// TIA Portal project "TESTV18" (V18)

(* hardware
DEVICE "Stazione S7-1500/ET200MP_1"  S7-1500 station
   slot 0: "Telaio di montaggio_0"  Rack  6ES7 590-1***0-0AA0
   slot 1: "PLC"  CPU 1511F-1 PN  6ES7 511-1FK02-0AB0  V2.8
      slot 3: "Display CPU_1"  6ES7591-1AA00-0AA0
      slot 32768: "Interfaccia PROFINET_1"  X1
         slot 32769: "Porta_1"  X1 P1
         slot 32770: "Porta_2"  X1 P2
      slot 34817: "Virtual CP interface port_1"  Virtual CP interface port  Virtual CP interface port
   slot 2: "AQ 4xU/I ST_1"  AQ 4xU/I ST  6ES7 532-5HD00-0AB0  V2.0
   slot 3: "AI 8xU/I HS_1"  AI 8xU/I HS  6ES7 531-7NF10-0AB0  V2.0
   slot 4: "DI 16x24VDC HF_1"  DI 16x24VDC HF  6ES7 521-1BH00-0AB0  V2.0
   slot 5: "DQ 16x24VDC/0.5A ST_1"  DQ 16x24VDC/0.5A ST  6ES7 522-1BH00-0AB0  V2.0
DEVICE "HMI"  TP700 Comfort
   slot 0: "HMI"  TP700 Comfort  6AV2 124-0GC01-0AX0  17.0.0.0
   slot 1: "HMI_RT_1"  TP700 Comfort  6AV2 124-0GC01-0AX0  17.0.0.0
   slot 5: "HMI.IE_CP_1"  PROFINET Interface  17.0.0.0
      slot 1: "Interfaccia_1 PROFINET"  PROFINET Interface
         slot 1: "Porta_1"  Port
         slot 2: "Porta_2"  Port
   slot 7: "HMI.MPI/DP_CP_1"  MPI/DP Interface  17.0.0.0
DEVICE "GSD device_1"  GSD.Device.PN
   slot 0: "Telaio di montaggio"  Rack  V1.0
   slot 0: "IAIPRT1"  RT Standard  IAI-PRT
      slot 0: "RT Standard"  RT Standard
      slot 1: "Interface"  Interface
         slot 1: "Port 1"  Port 1
   slot 1: "Input 1 word_1"  Input 1 word  IAI-PRT
      slot 0: "Input 1 word"  Input 1 word
   slot 2: "Input 1 word_2"  Input 1 word  IAI-PRT
      slot 0: "Input 1 word"  Input 1 word
   slot 3: "Input 1 word_3"  Input 1 word  IAI-PRT
      slot 0: "Input 1 word"  Input 1 word
   slot 4: "Input 1 word_4"  Input 1 word  IAI-PRT
      slot 0: "Input 1 word"  Input 1 word
   slot 5: "Input 1 word_5"  Input 1 word  IAI-PRT
      slot 0: "Input 1 word"  Input 1 word
   slot 6: "Input 1 word_6"  Input 1 word  IAI-PRT
      slot 0: "Input 1 word"  Input 1 word
   slot 7: "Input 1 word_7"  Input 1 word  IAI-PRT
      slot 0: "Input 1 word"  Input 1 word
   slot 8: "Input 1 word_8"  Input 1 word  IAI-PRT
      slot 0: "Input 1 word"  Input 1 word
   slot 9: "Input 1 word_9"  Input 1 word  IAI-PRT
      slot 0: "Input 1 word"  Input 1 word
   slot 10: "Input 1 word_10"  Input 1 word  IAI-PRT
      slot 0: "Input 1 word"  Input 1 word
   slot 11: "Input 1 word_11"  Input 1 word  IAI-PRT
      slot 0: "Input 1 word"  Input 1 word
   slot 12: "Input 1 word_12"  Input 1 word  IAI-PRT
      slot 0: "Input 1 word"  Input 1 word
   slot 13: "Input 1 word_13"  Input 1 word  IAI-PRT
      slot 0: "Input 1 word"  Input 1 word
   slot 14: "Input 1 word_14"  Input 1 word  IAI-PRT
      slot 0: "Input 1 word"  Input 1 word
   slot 15: "Input 1 word_15"  Input 1 word  IAI-PRT
      slot 0: "Input 1 word"  Input 1 word
   slot 16: "Input 1 word_16"  Input 1 word  IAI-PRT
      slot 0: "Input 1 word"  Input 1 word
   slot 17: "Output 1 word_1"  Output 1 word  IAI-PRT
      slot 0: "Output 1 word"  Output 1 word
   slot 18: "Output 1 word_2"  Output 1 word  IAI-PRT
      slot 0: "Output 1 word"  Output 1 word
   slot 19: "Output 1 word_3"  Output 1 word  IAI-PRT
      slot 0: "Output 1 word"  Output 1 word
   slot 20: "Output 1 word_4"  Output 1 word  IAI-PRT
      slot 0: "Output 1 word"  Output 1 word
   slot 21: "Output 1 word_5"  Output 1 word  IAI-PRT
      slot 0: "Output 1 word"  Output 1 word
   slot 22: "Output 1 word_6"  Output 1 word  IAI-PRT
      slot 0: "Output 1 word"  Output 1 word
   slot 23: "Output 1 word_7"  Output 1 word  IAI-PRT
      slot 0: "Output 1 word"  Output 1 word
   slot 24: "Output 1 word_8"  Output 1 word  IAI-PRT
      slot 0: "Output 1 word"  Output 1 word
   slot 25: "Output 1 word_9"  Output 1 word  IAI-PRT
      slot 0: "Output 1 word"  Output 1 word
   slot 26: "Output 1 word_10"  Output 1 word  IAI-PRT
      slot 0: "Output 1 word"  Output 1 word
   slot 27: "Output 1 word_11"  Output 1 word  IAI-PRT
      slot 0: "Output 1 word"  Output 1 word
   slot 28: "Output 1 word_12"  Output 1 word  IAI-PRT
      slot 0: "Output 1 word"  Output 1 word
   slot 29: "Output 1 word_13"  Output 1 word  IAI-PRT
      slot 0: "Output 1 word"  Output 1 word
   slot 30: "Output 1 word_14"  Output 1 word  IAI-PRT
      slot 0: "Output 1 word"  Output 1 word
   slot 31: "Output 1 word_15"  Output 1 word  IAI-PRT
      slot 0: "Output 1 word"  Output 1 word
   slot 32: "Output 1 word_16"  Output 1 word  IAI-PRT
      slot 0: "Output 1 word"  Output 1 word
*)

// ===== PLC "PLC"  CPU 1511F-1 PN =====

VAR_GLOBAL   // PLC tag table "Tabella delle variabili standard"
   "System_Byte" AT %MB16382 : Byte;
   "FirstScan" AT %M16382.0 : Bool;
   "DiagStatusUpdate" AT %M16382.1 : Bool;
   "AlwaysTRUE" AT %M16382.2 : Bool;
   "AlwaysFALSE" AT %M16382.3 : Bool;
   "Clock_Byte" AT %MB16383 : Byte;
   "Clock_10Hz" AT %M16383.0 : Bool;
   "Clock_5Hz" AT %M16383.1 : Bool;
   "Clock_2.5Hz" AT %M16383.2 : Bool;
   "Clock_2Hz" AT %M16383.3 : Bool;
   "Clock_1.25Hz" AT %M16383.4 : Bool;
   "Clock_1Hz" AT %M16383.5 : Bool;
   "Clock_0.625Hz" AT %M16383.6 : Bool;
   "Clock_0.5Hz" AT %M16383.7 : Bool;
   "Tag_1" AT %M0.0 : Bool;
   "Tag_2" AT %M0.1 : Bool;
   "Tag_3" AT %M0.3 : Bool;
   "Tag_4" AT %M0.4 : Bool;
   "Tag_5" AT %M0.5 : Bool;
   "Tag_6" AT %M0.6 : Bool;
   "Tag_7" AT %M0.7 : Bool;
   "Tag_8" AT %M500.0 : Bool;
   "Tag_9" AT %T100 : Timer;
   "Tag_10" AT %M0.2 : Bool;
   "Tag_11" AT %M2.0 : Bool;
   "Tag_12" AT %MD1000 : DWord;
   "Tag_13" AT %MW1000 : Word;
   "Tag_14" AT %MW1004 : UInt;
   "Tag_15" AT %Q2.0 : Bool;
   "Tag_16" AT %M5.0 : Bool;
   "Tag_17" AT %M5.1 : Bool;
   "Tag_18" AT %M5.2 : Bool;
   "Tag_19" AT %M5.3 : Bool;
   "Tag_20" AT %M4.0 : Bool;
   "Tag_21" AT %M4.1 : Bool;
   "Tag_22" AT %M3.0 : Bool;
   "Tag_23" AT %IW0 : Word;
   "Tag_24" AT %IB0 : Byte;
   "Tag_25" AT %IB16 : Byte;
   "Tag_26" AT %M2.1 : Bool;
   "Tag_27" AT %M2.3 : Bool;
   "Tag_28" AT %M2.4 : Bool;
   "Tag_29" AT %M2.5 : Bool;
   "Tag_30" AT %M2.6 : Bool;
   "Tag_31" AT %M2.7 : Bool;
   "Tag_32" AT %M2.2 : Bool;
   "Tag_33" AT %M3.1 : Bool;
   "Tag_34" AT %M3.2 : Bool;
   "Tag_35" AT %Q9.7 : Bool;
   "TGT_Pos" AT %QD10 : DWord;   // Position to be reached
   "Tag_37" AT %QD13 : DWord;
   "Tag_38" AT %QW10 : Word;
   "Tag_39" AT %QW11 : Word;
   "Tag_40" AT %QW13 : Word;
   "Tag_41" AT %QD12 : DWord;
   "Tag_42" AT %QD11 : DWord;
   "Tag_43" AT %QD34 : DWord;
   "CTRL_Sig2" AT %QD38 : DWord;   // Control dword signal 2
   "POS_BAND" AT %QD14 : DWord;   // Positioning band
   "SPE_mms" AT %QD18 : DWord;   // Speed mm/s
   "ZBO_ZBP" AT %QD22 : DWord;   // Zone boundary+
   "ZBO_ZBM" AT %QD26 : DWord;   // Zone boundary-
   "ACC_Accell" AT %QW30 : Word;   // Acceleration
   "DCL_Decell" AT %QW32 : Word;   // Deceleration
   "PLV_PressLimV" AT %QW34 : Word;   // Pressing current-limiting value
   "LCT_LoadCurrTh" AT %QW36 : Word;   // Load current threshold
   "Tag_36" AT %M1.0 : Bool;
   "Curr_POS" AT %ID18 : DWord;   // Current Position
   "Curr_CMD" AT %ID22 : DInt;   // Current command
   "Curr_SPD" AT %ID26 : UDInt;   // Current Speed
   "Allarm_COD" AT %ID30 : UDInt;   // Allarm Code
   "TotalMove_CNT" AT %ID38 : DInt;   // Total moving counter
   "TotalMove_DST" AT %ID42 : UDInt;   // Total moving distance
   "Status_DW" AT %ID46 : DWord;   // Status words PCON->PLC
END_VAR

TYPE "IAI_PCONPRTFM32OUT"
TITLE = IAI_PCONPRTFM32OUT
// Data type used for IAI PCON controller profinet configured in full mode (3 on parameter 84) with 32 word I/O occupied (0 on parameter 90)
   STRUCT
      Target_POS : DInt;   // Set the target position on the absolute coordinates.
      Positioning_BAND : UDInt;   // Positioning band
      Speed : UDInt;   // Specify the speed at which to move the actuator
      ZoneBNDP_BNDM : UDInt;   // The status signal PZONE turns ON when the current position is inside these +/- boundaries.
      Acceleration : USInt;   // Specify the acceleration at which to move the actuator
      Deceleration : USInt;   // Specify the deceleration at which to move the actuator
      Pressing_CLV : USInt;   // Specify the current- limiting value to be used during pressing operation.
      Load_current_threshold : USInt;   // Set the current threshold in this register when whether or not the load current exceeds the threshold is judged.
      CTRL1 : Struct   // Control WORD 1
         CTRL1_Sig_15 : Bool;   // Unavailable
         CTRL1_Sig_14 : Bool;   // Unavailable
         CTRL1_Sig_NTC1 : Bool;   // NTC1 (ACON only)
         CTRL1_Sig_NTC0 : Bool;   // NTC0 (ACON only)
         CTRL1_Sig_11 : Bool;   // Unavailable
         CTRL1_Sig_SMOD : Bool;   // SMOD (PCON only) Stopping control mode: When this signal is ON, servo control is performed during stopping.
         CTRL1_Sig_ASO1 : Bool;   // ASO1 Stop Mode 1 Select stop mode while standing
         CTRL1_Sig_ASO0 : Bool;   // ASO1 Stop Mode 0 Select stop mode while standing
         CTRL1_Sig_MOD1 : Bool;   // Acceleration / deceleration mode
         CTRL1_Sig_MOD0 : Bool;   // Acceleration / deceleration mode
         CTRL1_Sig_GSL1 : Bool;   // GSL1 (ACON only)
         CTRL1_Sig_GSL0 : Bool;   // GSL0 (ACON only)
         CTRL1_Sig_INC : Bool;   // Incremental Command: Absolute position commands are issued when this signal is OFF
         CTRL1_Sig_DIR : Bool;   // Pressing direction specification: “OFF” for the direction reducing the positioning band from the target position
         CTRL1_Sig_PUSH : Bool;   // Pressing specification : Positioning operation is performed when this signal is OFF
         CTRL1_Sig_00 : Bool;   // Unavailable
      END_STRUCT;
      CTRL2 : Struct   // Control WORD 2
         CTRL2_Sig_BKRL : Bool;   // Forced brake release: When it is turned ON, the brake is released
         CTRL2_Sig_RMOD : Bool;   // Operating mode selector : The AUTO mode is selected when this signal is OFF
         CTRL2_Sig_13 : Bool;   // Unavailable
         CTRL2_Sig_12 : Bool;   // Unavailable
         CTRL2_Sig_11 : Bool;   // Unavailable
         CTRL2_Sig_10 : Bool;   // Unavailable
         CTRL2_Sig_CLBR : Bool;   // Load cell calibration command (Dedicated for PCON-CBP/CGBP)
         "CTRL2_Sig_JOG+" : Bool;   // +Jog: “ON” for Movement in the Opposite Direction of Home
         "CTRL2_Sig_JOG-" : Bool;   // -Jog: “ON” for Movement in the Home Direction
         CTRL2_Sig_JVEL : Bool;   // Jog-speed/inch-distance switching
         CTRL2_Sig_JISL : Bool;   // Jog/inch switching: Jog operation is performed when this signal is OFF
         CTRL2_Sig_SON : Bool;   // GSL0 (ACON only)
         CTRL2_Sig_RES : Bool;   // Reset: A reset is performed when this signal turns ON.
         CTRL2_Sig_STP : Bool;   // Pause: A pause command is issued when this signal turns ON.
         CTRL2_Sig_HOME : Bool;   // Home return: A home-return command is issued when this signal turns ON.
         CTRL2_Sig_DSTR : Bool;   // Positioning start: A move command is issued when this signal turns ON.
      END_STRUCT;
   END_STRUCT;
END_TYPE

TYPE "IAI_PCONPRT"
   STRUCT
      PLCToPCON : "IAI_PCONPRTFM32OUT";
      PCONToPLC : "IAI_PCONPRTFM32IN";
   END_STRUCT;
END_TYPE

TYPE "IAI_PCONPRTFM32IN"
TITLE = IAI_PCONPRTFM32OUT
// Data type used for IAI PCON controller profinet configured in full mode (3 on parameter 84) with 32 word I/O occupied (0 on parameter 90)
   STRUCT
      Current_POS : DInt;   // Stores the current position. The unit is 0.01mm.
      Command_CUR : UDInt;   // Stores the currently commanded current. The unit is mA.
      Current_SPD : DInt;   // The current speed is indicated. The unit is 0.01mm/s. Positive value: The actuator is moving in the direction opposite home.
      Alarm_COD : UDInt;   // Stores an alarm code when an alarm (all alarms including message level ones) is generated.
      Current_LOA : DInt;   // Current load (Dedicated for PCON-CBP /CGBP)The unit is 0.01N.
      TotalMove_CNT : UDInt;   // Total moving conts (unit: times)
      TotalMove_DST : USInt;   // Total moving distance (unit: m)
      CTRL1 : Struct   // Control WORD 1
         STAT1_Sig_15 : Bool;   // Unavailable
         STAT1_Sig_14 : Bool;   // Unavailable
         STAT1_Sig_13 : Bool;   // Unavailable
         STAT1_Sig_12 : Bool;   // Unavailable
         STAT1_Sig_11 : Bool;   // Unavailable
         STAT1_Sig_10 : Bool;   // Unavailable
         STAT1_Sig_09 : Bool;   // Unavailable
         STAT1_Sig_08 : Bool;   // Unavailable
         STAT1_Sig_07 : Bool;   // Unavailable
         STAT1_Sig_06 : Bool;   // Unavailable
         STAT1_Sig_05 : Bool;   // Unavailable
         STAT1_Sig_04 : Bool;   // Unavailable
         STAT1_Sig_03 : Bool;   // Unavailable
         STAT1_Sig_02 : Bool;   // Unavailable
         CTRL1_Sig_CEND : Bool;   // Load cell calibration command. (Dedicated for PCON-CBP/CGBP)
         CTRL1_Sig_ALML : Bool;   // Light error status: Turns ON when light alarm (threshold exceeded for number of movement, etc.) that the operation can be continued with is issued. Note: ALM LED would not turn ON with a light error.
      END_STRUCT;
      CTRL2 : Struct   // Control WORD 2
         CTRL2_Sig_EMGS : Bool;   // Emergency stop: An emergency stop is actuated when this signal turns ON.
         CTRL2_Sig_PWR : Bool;   // Controller ready : This signal turns ON when the controller becomes ready.
         CTRL2_Sig_ZONE2 : Bool;   // Zone 2:“ON” for the current position within the zone set range
         CTRL2_Sig_ZONE1 : Bool;   // Zone 1:“ON” for the current position within the zone set range
         CTRL2_Sig_PZONE : Bool;   // Position zone: This signal turns ON when the current position is inside the specified position zone.
         CTRL2_Sig_LOAD : Bool;   // Load output judgment: When this signal is ON, the specified load has been reached.
         CTRL2_Sig_TRQS : Bool;   // Torque level: When this signal is ON, the specified load has been reached.
         CTRL2_Sig_RMDS : Bool;   // Operation mode status: This signal is OFF when the current mode is AUTO, or ON when the current mode is MANU.
         CTRL2_Sig_GHMS : Bool;   // Under Home return Operation: This signal remains ON while home return is in progress.
         CTRL2_Sig_PUSHS : Bool;   // Pressing in progress: This signal remains ON while pressing operation is in progress.
         CTRL2_Sig_PSFL : Bool;   // Pressing and a Miss: This signal turns ON when the actuator missed the work part in pressing operation.
         CTRL2_Sig_SV : Bool;   // Operation preparation end: This signal turns ON when the servo turns ON.
         CTRL2_Sig_ALM : Bool;   // Alarm: This signal turns ON when an alarm occurs.
         CTRL2_Sig_MOVE : Bool;   // Moving signal: This signal remains ON while the actuator is moving.
         CTRL2_Sig_HEND : Bool;   // Home return completion: This signal turns ON when home return is completed
         CTRL2_Sig_PEND : Bool;   // Positioning completion signal: This signal turns ON when positioning is completed.
      END_STRUCT;
   END_STRUCT;
END_TYPE

DATA_BLOCK "Main_Safety_RTG1_DB"   // DB1, F_DB
{ S7_Optimized_Access := 'TRUE' }
NAME : FUSI
VERSION : 0.1
// stored: InstanceOfName Main_Safety_RTG1
"Main_Safety_RTG1"
BEGIN
END_DATA_BLOCK

DATA_BLOCK "DB_AUX"   // DB3
{ S7_Optimized_Access := 'TRUE' }
VERSION : 0.1
   VAR
      FP : Array[0..10] of Bool;
      TARGET_POS : Array[0..4] of DInt;
      SPEED_POS : Array[0..4] of UDInt;
      ACC_DEC : USInt;
      AXIS1 : "IAI_PCONPRT";
      HMI_Bit : Struct
         HMIb1 : Bool;   // Load POS1
         HMIb2 : Bool;   // Load POS2
         HMIb3 : Bool;   // Load POS3
         HMIb4 : Bool;   // Load POS4
         HMIb5 : Bool;   // Servo ON
         HMIb6 : Bool;   // Start positioning
         HMIb7 : Bool;   // Homing
         HMIb8 : Bool;   // JOG+
         HMIb9 : Bool;   // JOG-
         HMIb10 : Bool;   // Reset allarm
         HMIb11 : Bool;
         HMIb12 : Bool;
         HMIb13 : Bool;
      END_STRUCT;
   END_VAR
BEGIN
END_DATA_BLOCK

FUNCTION_BLOCK "Main_Safety_RTG1"   // FB1, F_FBD
{ S7_Optimized_Access := 'TRUE' }
BEGIN
END_FUNCTION_BLOCK

ORGANIZATION_BLOCK "Main"   // OB1, LAD, ProgramCycle
TITLE = "Main Program Sweep (Cycle)"
{ S7_Optimized_Access := 'TRUE' }
VERSION : 0.1
   VAR_INPUT
      Initial_Call : Bool;   // Initial call of this OB
      Remanence : Bool;   // =True, if remanent data are available
   END_VAR
BEGIN

REGION Network 1: IAI controllers side input register PLC -> PCON
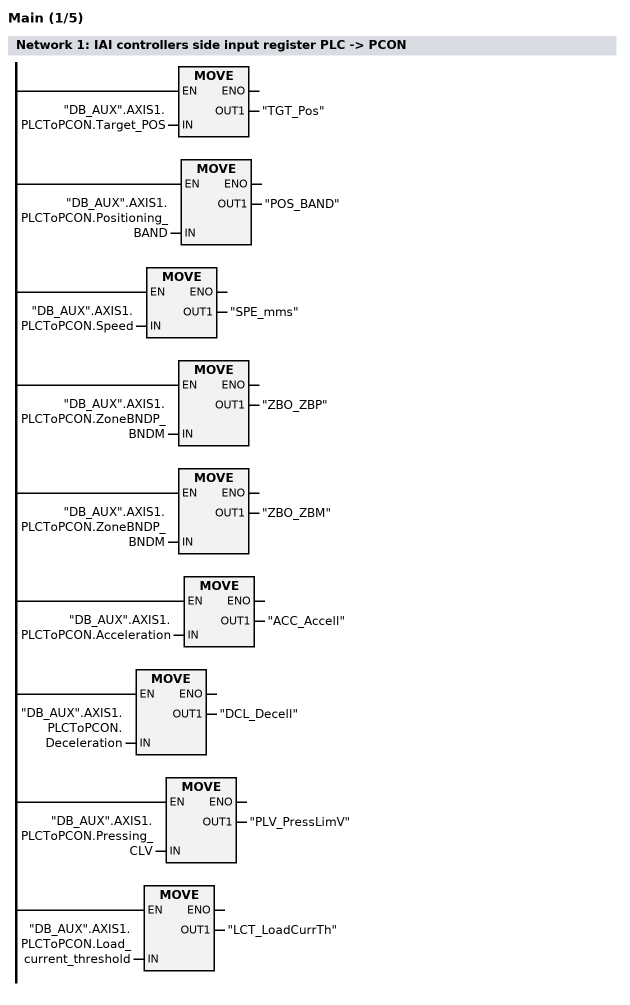
   RUNG wire#powerrail
      Move(in := "DB_AUX".AXIS1.PLCToPCON.Target_POS, out1 => "TGT_Pos")
   END_RUNG
   RUNG wire#powerrail
      Move(in := "DB_AUX".AXIS1.PLCToPCON.Positioning_BAND, out1 => "POS_BAND")
   END_RUNG
   RUNG wire#powerrail
      Move(in := "DB_AUX".AXIS1.PLCToPCON.Speed, out1 => "SPE_mms")
   END_RUNG
   RUNG wire#powerrail
      Move(in := "DB_AUX".AXIS1.PLCToPCON.ZoneBNDP_BNDM, out1 => "ZBO_ZBP")
   END_RUNG
   RUNG wire#powerrail
      Move(in := "DB_AUX".AXIS1.PLCToPCON.ZoneBNDP_BNDM, out1 => "ZBO_ZBM")
   END_RUNG
   RUNG wire#powerrail
      Move(in := "DB_AUX".AXIS1.PLCToPCON.Acceleration, out1 => "ACC_Accell")
   END_RUNG
   RUNG wire#powerrail
      Move(in := "DB_AUX".AXIS1.PLCToPCON.Deceleration, out1 => "DCL_Decell")
   END_RUNG
   RUNG wire#powerrail
      Move(in := "DB_AUX".AXIS1.PLCToPCON.Pressing_CLV, out1 => "PLV_PressLimV")
   END_RUNG
   RUNG wire#powerrail
      Move(in := "DB_AUX".AXIS1.PLCToPCON.Load_current_threshold, out1 => "LCT_LoadCurrTh")
   END_RUNG
   // the same network as SCL:
   "TGT_Pos" := "DB_AUX".AXIS1.PLCToPCON.Target_POS;
   "POS_BAND" := "DB_AUX".AXIS1.PLCToPCON.Positioning_BAND;
   "SPE_mms" := "DB_AUX".AXIS1.PLCToPCON.Speed;
   "ZBO_ZBP" := "DB_AUX".AXIS1.PLCToPCON.ZoneBNDP_BNDM;
   "ZBO_ZBM" := "DB_AUX".AXIS1.PLCToPCON.ZoneBNDP_BNDM;
   "ACC_Accell" := "DB_AUX".AXIS1.PLCToPCON.Acceleration;
   "DCL_Decell" := "DB_AUX".AXIS1.PLCToPCON.Deceleration;
   "PLV_PressLimV" := "DB_AUX".AXIS1.PLCToPCON.Pressing_CLV;
   "LCT_LoadCurrTh" := "DB_AUX".AXIS1.PLCToPCON.Load_current_threshold;
END_REGION

REGION Network 2: IAI controllers side input register PLC -> PCON
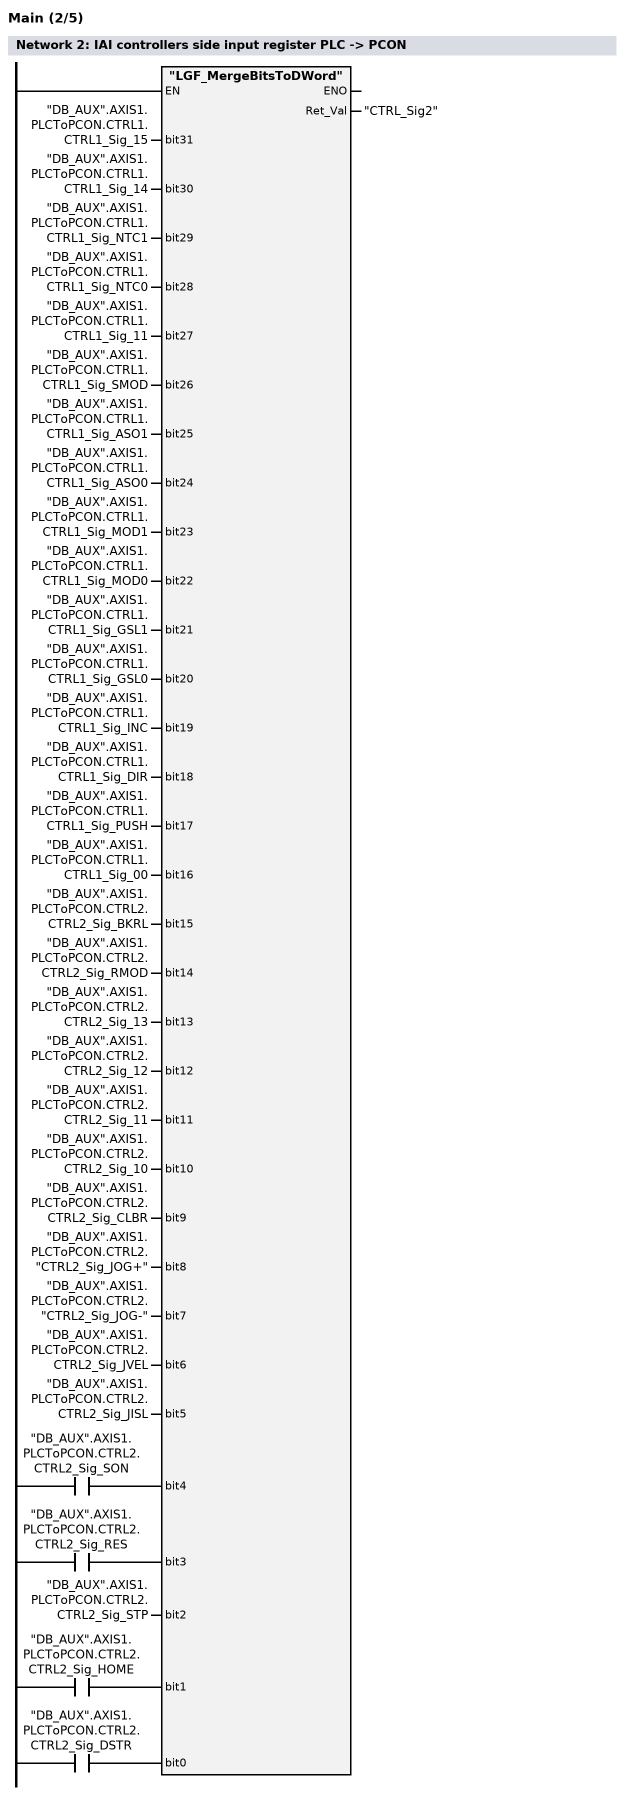
   RUNG wire#powerrail
      "LGF_MergeBitsToDWord"(bit4 := wire#w1, bit3 := wire#w2, bit1 := wire#w3, bit0 := wire#w4, bit31 := "DB_AUX".AXIS1.PLCToPCON.CTRL1.CTRL1_Sig_15, bit30 := "DB_AUX".AXIS1.PLCToPCON.CTRL1.CTRL1_Sig_14, bit29 := "DB_AUX".AXIS1.PLCToPCON.CTRL1.CTRL1_Sig_NTC1, bit28 := "DB_AUX".AXIS1.PLCToPCON.CTRL1.CTRL1_Sig_NTC0, bit27 := "DB_AUX".AXIS1.PLCToPCON.CTRL1.CTRL1_Sig_11, bit26 := "DB_AUX".AXIS1.PLCToPCON.CTRL1.CTRL1_Sig_SMOD, bit25 := "DB_AUX".AXIS1.PLCToPCON.CTRL1.CTRL1_Sig_ASO1, bit24 := "DB_AUX".AXIS1.PLCToPCON.CTRL1.CTRL1_Sig_ASO0, bit23 := "DB_AUX".AXIS1.PLCToPCON.CTRL1.CTRL1_Sig_MOD1, bit22 := "DB_AUX".AXIS1.PLCToPCON.CTRL1.CTRL1_Sig_MOD0, bit21 := "DB_AUX".AXIS1.PLCToPCON.CTRL1.CTRL1_Sig_GSL1, bit20 := "DB_AUX".AXIS1.PLCToPCON.CTRL1.CTRL1_Sig_GSL0, bit19 := "DB_AUX".AXIS1.PLCToPCON.CTRL1.CTRL1_Sig_INC, bit18 := "DB_AUX".AXIS1.PLCToPCON.CTRL1.CTRL1_Sig_DIR, bit17 := "DB_AUX".AXIS1.PLCToPCON.CTRL1.CTRL1_Sig_PUSH, bit16 := "DB_AUX".AXIS1.PLCToPCON.CTRL1.CTRL1_Sig_00, bit15 := "DB_AUX".AXIS1.PLCToPCON.CTRL2.CTRL2_Sig_BKRL, bit14 := "DB_AUX".AXIS1.PLCToPCON.CTRL2.CTRL2_Sig_RMOD, bit13 := "DB_AUX".AXIS1.PLCToPCON.CTRL2.CTRL2_Sig_13, bit12 := "DB_AUX".AXIS1.PLCToPCON.CTRL2.CTRL2_Sig_12, bit11 := "DB_AUX".AXIS1.PLCToPCON.CTRL2.CTRL2_Sig_11, bit10 := "DB_AUX".AXIS1.PLCToPCON.CTRL2.CTRL2_Sig_10, bit9 := "DB_AUX".AXIS1.PLCToPCON.CTRL2.CTRL2_Sig_CLBR, bit8 := "DB_AUX".AXIS1.PLCToPCON.CTRL2."CTRL2_Sig_JOG+", bit7 := "DB_AUX".AXIS1.PLCToPCON.CTRL2."CTRL2_Sig_JOG-", bit6 := "DB_AUX".AXIS1.PLCToPCON.CTRL2.CTRL2_Sig_JVEL, bit5 := "DB_AUX".AXIS1.PLCToPCON.CTRL2.CTRL2_Sig_JISL, bit2 := "DB_AUX".AXIS1.PLCToPCON.CTRL2.CTRL2_Sig_STP, Ret_Val => "CTRL_Sig2")
   END_RUNG
   RUNG wire#powerrail
      Contact( "DB_AUX".AXIS1.PLCToPCON.CTRL2.CTRL2_Sig_SON )
   END_RUNG wire#w1
   RUNG wire#powerrail
      Contact( "DB_AUX".AXIS1.PLCToPCON.CTRL2.CTRL2_Sig_RES )
   END_RUNG wire#w2
   RUNG wire#powerrail
      Contact( "DB_AUX".AXIS1.PLCToPCON.CTRL2.CTRL2_Sig_HOME )
   END_RUNG wire#w3
   RUNG wire#powerrail
      Contact( "DB_AUX".AXIS1.PLCToPCON.CTRL2.CTRL2_Sig_DSTR )
   END_RUNG wire#w4
   // the same network as SCL:
   "CTRL_Sig2" := "LGF_MergeBitsToDWord"(bit31 := "DB_AUX".AXIS1.PLCToPCON.CTRL1.CTRL1_Sig_15,
                           bit30 := "DB_AUX".AXIS1.PLCToPCON.CTRL1.CTRL1_Sig_14,
                           bit29 := "DB_AUX".AXIS1.PLCToPCON.CTRL1.CTRL1_Sig_NTC1,
                           bit28 := "DB_AUX".AXIS1.PLCToPCON.CTRL1.CTRL1_Sig_NTC0,
                           bit27 := "DB_AUX".AXIS1.PLCToPCON.CTRL1.CTRL1_Sig_11,
                           bit26 := "DB_AUX".AXIS1.PLCToPCON.CTRL1.CTRL1_Sig_SMOD,
                           bit25 := "DB_AUX".AXIS1.PLCToPCON.CTRL1.CTRL1_Sig_ASO1,
                           bit24 := "DB_AUX".AXIS1.PLCToPCON.CTRL1.CTRL1_Sig_ASO0,
                           bit23 := "DB_AUX".AXIS1.PLCToPCON.CTRL1.CTRL1_Sig_MOD1,
                           bit22 := "DB_AUX".AXIS1.PLCToPCON.CTRL1.CTRL1_Sig_MOD0,
                           bit21 := "DB_AUX".AXIS1.PLCToPCON.CTRL1.CTRL1_Sig_GSL1,
                           bit20 := "DB_AUX".AXIS1.PLCToPCON.CTRL1.CTRL1_Sig_GSL0,
                           bit19 := "DB_AUX".AXIS1.PLCToPCON.CTRL1.CTRL1_Sig_INC,
                           bit18 := "DB_AUX".AXIS1.PLCToPCON.CTRL1.CTRL1_Sig_DIR,
                           bit17 := "DB_AUX".AXIS1.PLCToPCON.CTRL1.CTRL1_Sig_PUSH,
                           bit16 := "DB_AUX".AXIS1.PLCToPCON.CTRL1.CTRL1_Sig_00,
                           bit15 := "DB_AUX".AXIS1.PLCToPCON.CTRL2.CTRL2_Sig_BKRL,
                           bit14 := "DB_AUX".AXIS1.PLCToPCON.CTRL2.CTRL2_Sig_RMOD,
                           bit13 := "DB_AUX".AXIS1.PLCToPCON.CTRL2.CTRL2_Sig_13,
                           bit12 := "DB_AUX".AXIS1.PLCToPCON.CTRL2.CTRL2_Sig_12,
                           bit11 := "DB_AUX".AXIS1.PLCToPCON.CTRL2.CTRL2_Sig_11,
                           bit10 := "DB_AUX".AXIS1.PLCToPCON.CTRL2.CTRL2_Sig_10,
                           bit9 := "DB_AUX".AXIS1.PLCToPCON.CTRL2.CTRL2_Sig_CLBR,
                           bit8 := "DB_AUX".AXIS1.PLCToPCON.CTRL2."CTRL2_Sig_JOG+",
                           bit7 := "DB_AUX".AXIS1.PLCToPCON.CTRL2."CTRL2_Sig_JOG-",
                           bit6 := "DB_AUX".AXIS1.PLCToPCON.CTRL2.CTRL2_Sig_JVEL,
                           bit5 := "DB_AUX".AXIS1.PLCToPCON.CTRL2.CTRL2_Sig_JISL,
                           bit4 := "DB_AUX".AXIS1.PLCToPCON.CTRL2.CTRL2_Sig_SON,
                           bit3 := "DB_AUX".AXIS1.PLCToPCON.CTRL2.CTRL2_Sig_RES,
                           bit2 := "DB_AUX".AXIS1.PLCToPCON.CTRL2.CTRL2_Sig_STP,
                           bit1 := "DB_AUX".AXIS1.PLCToPCON.CTRL2.CTRL2_Sig_HOME,
                           bit0 := "DB_AUX".AXIS1.PLCToPCON.CTRL2.CTRL2_Sig_DSTR);
END_REGION

REGION Network 3: --------------------------------------------------------------------------------
END_REGION

REGION Network 4: IAI controllers side input register PCON->PLC
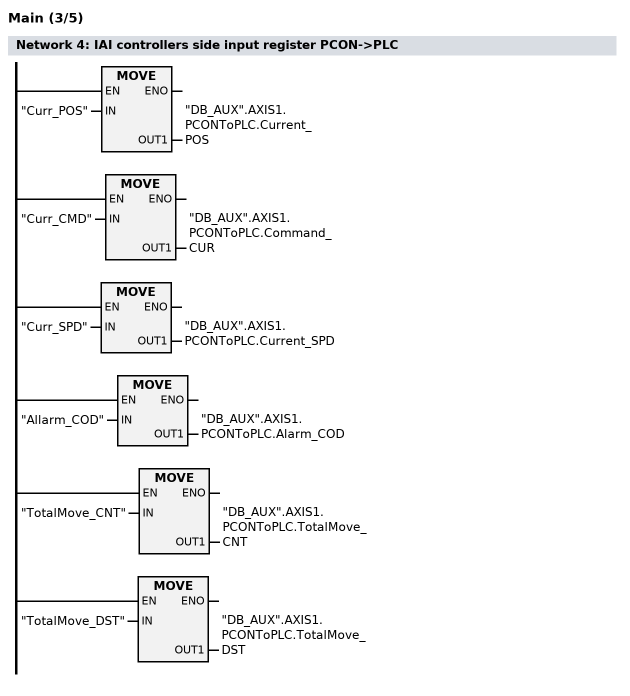
   RUNG wire#powerrail
      Move(in := "Curr_POS", out1 => "DB_AUX".AXIS1.PCONToPLC.Current_POS)
   END_RUNG
   RUNG wire#powerrail
      Move(in := "Curr_CMD", out1 => "DB_AUX".AXIS1.PCONToPLC.Command_CUR)
   END_RUNG
   RUNG wire#powerrail
      Move(in := "Curr_SPD", out1 => "DB_AUX".AXIS1.PCONToPLC.Current_SPD)
   END_RUNG
   RUNG wire#powerrail
      Move(in := "Allarm_COD", out1 => "DB_AUX".AXIS1.PCONToPLC.Alarm_COD)
   END_RUNG
   RUNG wire#powerrail
      Move(in := "TotalMove_CNT", out1 => "DB_AUX".AXIS1.PCONToPLC.TotalMove_CNT)
   END_RUNG
   RUNG wire#powerrail
      Move(in := "TotalMove_DST", out1 => "DB_AUX".AXIS1.PCONToPLC.TotalMove_DST)
   END_RUNG
   // the same network as SCL:
   "DB_AUX".AXIS1.PCONToPLC.Current_POS := "Curr_POS";
   "DB_AUX".AXIS1.PCONToPLC.Command_CUR := "Curr_CMD";
   "DB_AUX".AXIS1.PCONToPLC.Current_SPD := "Curr_SPD";
   "DB_AUX".AXIS1.PCONToPLC.Alarm_COD := "Allarm_COD";
   "DB_AUX".AXIS1.PCONToPLC.TotalMove_CNT := "TotalMove_CNT";
   "DB_AUX".AXIS1.PCONToPLC.TotalMove_DST := "TotalMove_DST";
END_REGION

REGION Network 5: IAI controllers side input register PCON->PLC
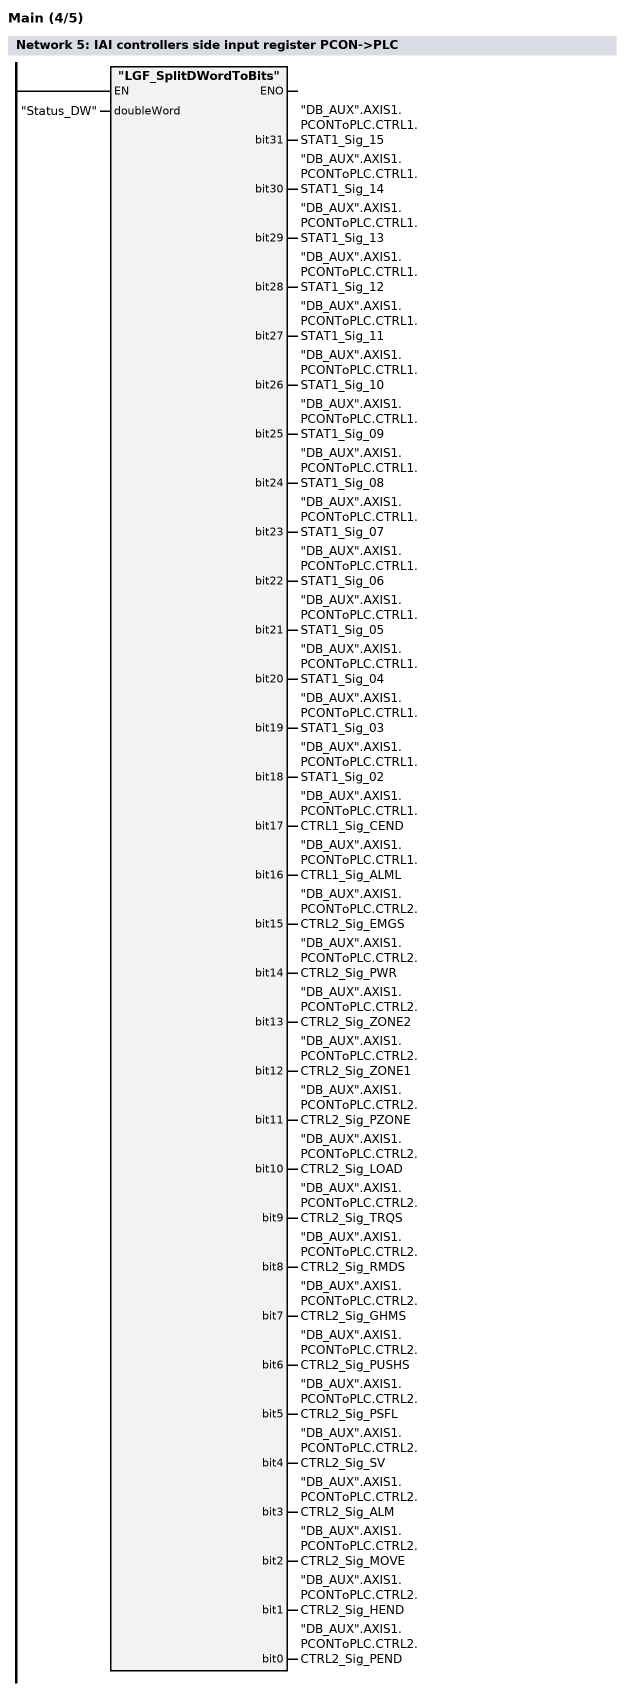
   RUNG wire#powerrail
      "LGF_SplitDWordToBits"(doubleWord := "Status_DW", bit31 => "DB_AUX".AXIS1.PCONToPLC.CTRL1.STAT1_Sig_15, bit30 => "DB_AUX".AXIS1.PCONToPLC.CTRL1.STAT1_Sig_14, bit29 => "DB_AUX".AXIS1.PCONToPLC.CTRL1.STAT1_Sig_13, bit28 => "DB_AUX".AXIS1.PCONToPLC.CTRL1.STAT1_Sig_12, bit27 => "DB_AUX".AXIS1.PCONToPLC.CTRL1.STAT1_Sig_11, bit26 => "DB_AUX".AXIS1.PCONToPLC.CTRL1.STAT1_Sig_10, bit25 => "DB_AUX".AXIS1.PCONToPLC.CTRL1.STAT1_Sig_09, bit24 => "DB_AUX".AXIS1.PCONToPLC.CTRL1.STAT1_Sig_08, bit23 => "DB_AUX".AXIS1.PCONToPLC.CTRL1.STAT1_Sig_07, bit22 => "DB_AUX".AXIS1.PCONToPLC.CTRL1.STAT1_Sig_06, bit21 => "DB_AUX".AXIS1.PCONToPLC.CTRL1.STAT1_Sig_05, bit20 => "DB_AUX".AXIS1.PCONToPLC.CTRL1.STAT1_Sig_04, bit19 => "DB_AUX".AXIS1.PCONToPLC.CTRL1.STAT1_Sig_03, bit18 => "DB_AUX".AXIS1.PCONToPLC.CTRL1.STAT1_Sig_02, bit17 => "DB_AUX".AXIS1.PCONToPLC.CTRL1.CTRL1_Sig_CEND, bit16 => "DB_AUX".AXIS1.PCONToPLC.CTRL1.CTRL1_Sig_ALML, bit15 => "DB_AUX".AXIS1.PCONToPLC.CTRL2.CTRL2_Sig_EMGS, bit14 => "DB_AUX".AXIS1.PCONToPLC.CTRL2.CTRL2_Sig_PWR, bit13 => "DB_AUX".AXIS1.PCONToPLC.CTRL2.CTRL2_Sig_ZONE2, bit12 => "DB_AUX".AXIS1.PCONToPLC.CTRL2.CTRL2_Sig_ZONE1, bit11 => "DB_AUX".AXIS1.PCONToPLC.CTRL2.CTRL2_Sig_PZONE, bit10 => "DB_AUX".AXIS1.PCONToPLC.CTRL2.CTRL2_Sig_LOAD, bit9 => "DB_AUX".AXIS1.PCONToPLC.CTRL2.CTRL2_Sig_TRQS, bit8 => "DB_AUX".AXIS1.PCONToPLC.CTRL2.CTRL2_Sig_RMDS, bit7 => "DB_AUX".AXIS1.PCONToPLC.CTRL2.CTRL2_Sig_GHMS, bit6 => "DB_AUX".AXIS1.PCONToPLC.CTRL2.CTRL2_Sig_PUSHS, bit5 => "DB_AUX".AXIS1.PCONToPLC.CTRL2.CTRL2_Sig_PSFL, bit4 => "DB_AUX".AXIS1.PCONToPLC.CTRL2.CTRL2_Sig_SV, bit3 => "DB_AUX".AXIS1.PCONToPLC.CTRL2.CTRL2_Sig_ALM, bit2 => "DB_AUX".AXIS1.PCONToPLC.CTRL2.CTRL2_Sig_MOVE, bit1 => "DB_AUX".AXIS1.PCONToPLC.CTRL2.CTRL2_Sig_HEND, bit0 => "DB_AUX".AXIS1.PCONToPLC.CTRL2.CTRL2_Sig_PEND)
   END_RUNG
   // the same network as SCL:
   "LGF_SplitDWordToBits"(doubleWord := "Status_DW",
                          bit31 => "DB_AUX".AXIS1.PCONToPLC.CTRL1.STAT1_Sig_15,
                          bit30 => "DB_AUX".AXIS1.PCONToPLC.CTRL1.STAT1_Sig_14,
                          bit29 => "DB_AUX".AXIS1.PCONToPLC.CTRL1.STAT1_Sig_13,
                          bit28 => "DB_AUX".AXIS1.PCONToPLC.CTRL1.STAT1_Sig_12,
                          bit27 => "DB_AUX".AXIS1.PCONToPLC.CTRL1.STAT1_Sig_11,
                          bit26 => "DB_AUX".AXIS1.PCONToPLC.CTRL1.STAT1_Sig_10,
                          bit25 => "DB_AUX".AXIS1.PCONToPLC.CTRL1.STAT1_Sig_09,
                          bit24 => "DB_AUX".AXIS1.PCONToPLC.CTRL1.STAT1_Sig_08,
                          bit23 => "DB_AUX".AXIS1.PCONToPLC.CTRL1.STAT1_Sig_07,
                          bit22 => "DB_AUX".AXIS1.PCONToPLC.CTRL1.STAT1_Sig_06,
                          bit21 => "DB_AUX".AXIS1.PCONToPLC.CTRL1.STAT1_Sig_05,
                          bit20 => "DB_AUX".AXIS1.PCONToPLC.CTRL1.STAT1_Sig_04,
                          bit19 => "DB_AUX".AXIS1.PCONToPLC.CTRL1.STAT1_Sig_03,
                          bit18 => "DB_AUX".AXIS1.PCONToPLC.CTRL1.STAT1_Sig_02,
                          bit17 => "DB_AUX".AXIS1.PCONToPLC.CTRL1.CTRL1_Sig_CEND,
                          bit16 => "DB_AUX".AXIS1.PCONToPLC.CTRL1.CTRL1_Sig_ALML,
                          bit15 => "DB_AUX".AXIS1.PCONToPLC.CTRL2.CTRL2_Sig_EMGS,
                          bit14 => "DB_AUX".AXIS1.PCONToPLC.CTRL2.CTRL2_Sig_PWR,
                          bit13 => "DB_AUX".AXIS1.PCONToPLC.CTRL2.CTRL2_Sig_ZONE2,
                          bit12 => "DB_AUX".AXIS1.PCONToPLC.CTRL2.CTRL2_Sig_ZONE1,
                          bit11 => "DB_AUX".AXIS1.PCONToPLC.CTRL2.CTRL2_Sig_PZONE,
                          bit10 => "DB_AUX".AXIS1.PCONToPLC.CTRL2.CTRL2_Sig_LOAD,
                          bit9 => "DB_AUX".AXIS1.PCONToPLC.CTRL2.CTRL2_Sig_TRQS,
                          bit8 => "DB_AUX".AXIS1.PCONToPLC.CTRL2.CTRL2_Sig_RMDS,
                          bit7 => "DB_AUX".AXIS1.PCONToPLC.CTRL2.CTRL2_Sig_GHMS,
                          bit6 => "DB_AUX".AXIS1.PCONToPLC.CTRL2.CTRL2_Sig_PUSHS,
                          bit5 => "DB_AUX".AXIS1.PCONToPLC.CTRL2.CTRL2_Sig_PSFL,
                          bit4 => "DB_AUX".AXIS1.PCONToPLC.CTRL2.CTRL2_Sig_SV,
                          bit3 => "DB_AUX".AXIS1.PCONToPLC.CTRL2.CTRL2_Sig_ALM,
                          bit2 => "DB_AUX".AXIS1.PCONToPLC.CTRL2.CTRL2_Sig_MOVE,
                          bit1 => "DB_AUX".AXIS1.PCONToPLC.CTRL2.CTRL2_Sig_HEND,
                          bit0 => "DB_AUX".AXIS1.PCONToPLC.CTRL2.CTRL2_Sig_PEND);
END_REGION

REGION Network 6: --------------------------------------------------------------------------------
END_REGION

REGION Network 7: HMI Interface
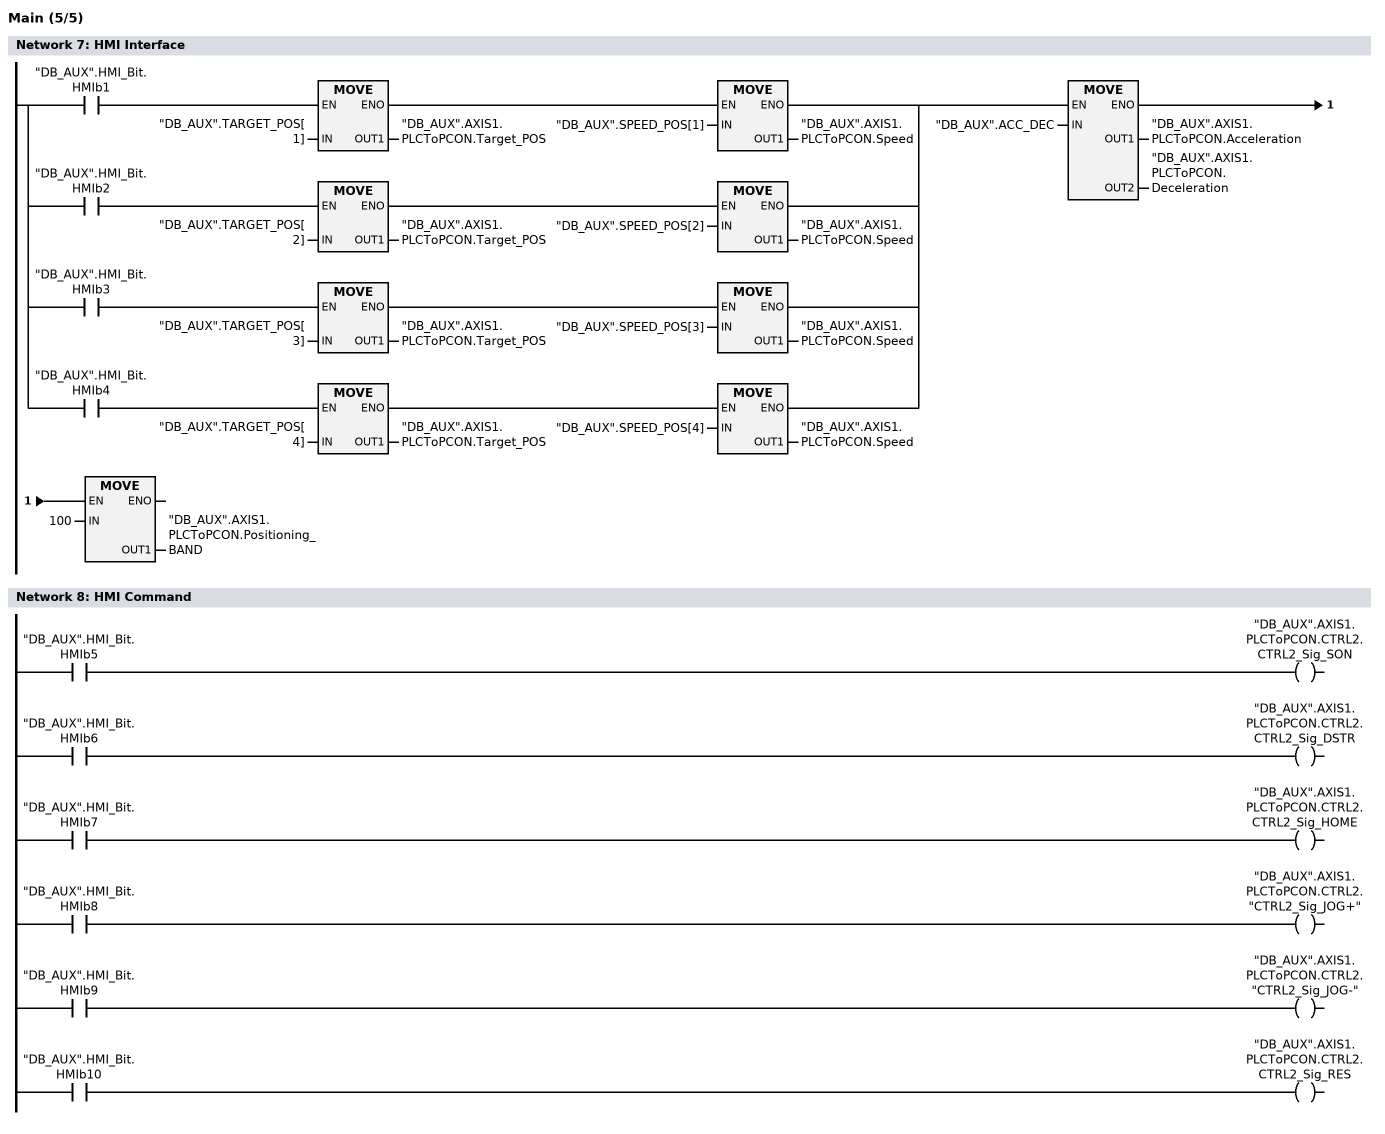
   RUNG wire#powerrail
      Contact( "DB_AUX".HMI_Bit.HMIb1 )
      Move(in := "DB_AUX".TARGET_POS[1], out1 => "DB_AUX".AXIS1.PLCToPCON.Target_POS)
      Move(in := "DB_AUX".SPEED_POS[1], out1 => "DB_AUX".AXIS1.PLCToPCON.Speed)
      wire#w1
      Move(in := "DB_AUX".ACC_DEC, out1 => "DB_AUX".AXIS1.PLCToPCON.Acceleration, out2 => "DB_AUX".AXIS1.PLCToPCON.Deceleration)
      Move(in := 100, out1 => "DB_AUX".AXIS1.PLCToPCON.Positioning_BAND)
   END_RUNG
   RUNG wire#powerrail
      Contact( "DB_AUX".HMI_Bit.HMIb2 )
      Move(in := "DB_AUX".TARGET_POS[2], out1 => "DB_AUX".AXIS1.PLCToPCON.Target_POS)
      Move(in := "DB_AUX".SPEED_POS[2], out1 => "DB_AUX".AXIS1.PLCToPCON.Speed)
   END_RUNG wire#w1
   RUNG wire#powerrail
      Contact( "DB_AUX".HMI_Bit.HMIb3 )
      Move(in := "DB_AUX".TARGET_POS[3], out1 => "DB_AUX".AXIS1.PLCToPCON.Target_POS)
      Move(in := "DB_AUX".SPEED_POS[3], out1 => "DB_AUX".AXIS1.PLCToPCON.Speed)
   END_RUNG wire#w1
   RUNG wire#powerrail
      Contact( "DB_AUX".HMI_Bit.HMIb4 )
      Move(in := "DB_AUX".TARGET_POS[4], out1 => "DB_AUX".AXIS1.PLCToPCON.Target_POS)
      Move(in := "DB_AUX".SPEED_POS[4], out1 => "DB_AUX".AXIS1.PLCToPCON.Speed)
   END_RUNG wire#w1
   // the same network as SCL:
   IF "DB_AUX".HMI_Bit.HMIb1 THEN
       "DB_AUX".AXIS1.PLCToPCON.Target_POS := "DB_AUX".TARGET_POS[1];
       "DB_AUX".AXIS1.PLCToPCON.Speed := "DB_AUX".SPEED_POS[1];
   END_IF;
   IF "DB_AUX".HMI_Bit.HMIb2 THEN
       "DB_AUX".AXIS1.PLCToPCON.Target_POS := "DB_AUX".TARGET_POS[2];
       "DB_AUX".AXIS1.PLCToPCON.Speed := "DB_AUX".SPEED_POS[2];
   END_IF;
   IF "DB_AUX".HMI_Bit.HMIb3 THEN
       "DB_AUX".AXIS1.PLCToPCON.Target_POS := "DB_AUX".TARGET_POS[3];
       "DB_AUX".AXIS1.PLCToPCON.Speed := "DB_AUX".SPEED_POS[3];
   END_IF;
   IF "DB_AUX".HMI_Bit.HMIb4 THEN
       "DB_AUX".AXIS1.PLCToPCON.Target_POS := "DB_AUX".TARGET_POS[4];
       "DB_AUX".AXIS1.PLCToPCON.Speed := "DB_AUX".SPEED_POS[4];
   END_IF;
   IF "DB_AUX".HMI_Bit.HMIb1 OR "DB_AUX".HMI_Bit.HMIb2 OR "DB_AUX".HMI_Bit.HMIb3 OR "DB_AUX".HMI_Bit.HMIb4 THEN
       "DB_AUX".AXIS1.PLCToPCON.Acceleration := "DB_AUX".ACC_DEC;
       "DB_AUX".AXIS1.PLCToPCON.Deceleration := "DB_AUX".ACC_DEC;
       "DB_AUX".AXIS1.PLCToPCON.Positioning_BAND := 100;
   END_IF;
END_REGION
